screen "MTA-TiemposCmpAlta" 1280x800, template "Plantilla"
   TextField "Campo de texto_3" at 278,160 size 235x27; Text 'Tiempo apagado Sopladora'
   IOField "Campo ES_5" at 889,160 size 90x23; FormatPattern 99; Unit  min
      ProcessValue <- "TiempoSop"
   TextField "Campo de texto_1" at 278,288 size 268x27; Text 'Tiempo de compresor en vacío'
   IOField "Campo ES_1" at 889,288 size 90x23; FormatPattern 99; Unit  min
      ProcessValue <- "TiempoenVacío"
   TextField "Campo de texto_2" at 278,432 size 339x27; Text 'Tiempo sin requerimiento de compresor'
   IOField "Campo ES_2" at 889,432 size 90x23; FormatPattern 99; Unit  min
      ProcessValue <- "TiemposinReq"
   TextField "Campo de texto_4" at 286,192 size 586x36; Text 'Una vez deshabilitada una sopladora, los requisitos de marcha de compresores se mantienen durante éste tiempo.'
   TextField "Campo de texto_5" at 286,320 size 616x52; Text 'Es el tiempo máximo durante el cual el compresor quedará funcionando en vacío. Una vez cumplido éste tiempo, el compresor será pasará al estado de "sin requerimiento". Si el compresor vuelve a ser requerido en carga, se pondrá en marcha sin requerir intervención del usuario'
   TextField "Campo de texto_6" at 286,464 size 578x36; Text 'Transcurrido éste tiempo en el estado “Sin requerimiento”, pasará al estado “sin marcha”, donde sí requerirá que se pulse el botón de MARCHA en caso de ser necesitado.'
   Button "Botón_12" at 1105,638 size 160x49; TextOff 'Volver'
      on Click: function_efd93a16()
   TextField "Campo de texto_7" at 477,9 size 326x27; Text 'Configuración de Tiempos Alta presión'

screen "MTA-TorresCAV" 1280x800, template "Plantilla"
   GraphicView "Visor de gráficos_9" at 71,137 size 234x255; Picture "torreFINAL4_1"
   GraphicView "Visor de gráficos_11" at 71,137 size 234x255; Picture "torreFINAL4B_1"
   GraphicView "Visor de gráficos_14" at 71,137 size 234x255; Picture "torreFINAL4C_1"
      Visibility <- "BombaTorreON2"
   GraphicView "Visor de gráficos_1" at 271,121 size 282x311; Picture "torreFINAL4_1"
   GraphicView "Visor de gráficos_2" at 271,121 size 282x311; Picture "torreFINAL4B_1"
   GraphicView "Visor de gráficos_3" at 271,121 size 282x311; Picture "torreFINAL4C_1"
      Visibility <- "BombaTorreON2"
   Polygon "Polígono_2" at 106,411 size 18x54
      Appearance <- "FT1_AGUA"
   ScreenModuleView "Faceplate_9_2" at 831,282 size 221x68
      Guid_{11997190-23979} <- "HabilitaciónMV030"
      Guid_{11997190-23983} <- "ParadaMV030"
      Guid_{11997190-23981} <- "MarchaMV030"
      Guid_{11997190-23989} <- "SP-OFF-V030"
      Guid_{11997190-23976} <- "DeshabilitaciónMV030"
      Guid_{11997190-23987} <- "SP-ON-V030"
      Guid_{11997190-23985} <- "MenuV030"
   ScreenModuleView "Faceplate_9_1" at 831,173 size 221x68
      Guid_{11997190-23979} <- "HabilitaciónMV031"
      Guid_{11997190-23983} <- "ParadaMV031"
      Guid_{11997190-23981} <- "MarchaMV031"
      Guid_{11997190-23989} <- "SP-OFF-V031"
      Guid_{11997190-23976} <- "DeshabilitaciónMV031"
      Guid_{11997190-23987} <- "SP-ON-V031"
      Guid_{11997190-23985} <- "MenuV031"
   Polygon "Polígono_4" at 60,416 size 46x49
      Appearance <- "FT1_AGUA"
   GraphicView "Visor de gráficos_17" at 7,412 size 77x78; Picture "tuboXXX5_1"
   GraphicView "Visor de gráficos_16" at 340,421 size 190x41; Picture "tuboXXX4"
   TextField "Campo de texto_23" at 647,286 size 126x32; Text 'Ventilador 2'
   TextField "Campo de texto_3" at 647,178 size 126x32; Text 'Ventilador 1'
   GraphicIOField "Campo ES gráfico_4" at 638,358 size 511x6; PictureList "Indicador"
      ProcessValue <- "AnimaMV030"
   GraphicIOField "Campo ES gráfico_5" at 638,250 size 511x6; PictureList "Indicador"
      ProcessValue <- "AnimaMV031"
   SymbolicIOField "Campo ES simbólico_6" at 649,322 size 170x21; TextOff '0'; TextOn '1'; TextList "EstadoMotor"
      ProcessValue <- "AnimaMV030"
   SymbolicIOField "Campo ES simbólico_2" at 649,214 size 170x21; TextOff '0'; TextOn '1'; TextList "EstadoMotor"
      ProcessValue <- "AnimaMV031"
   Switch "Interruptor_5" at 782,288 size 29x29; TextOn '1'; TextOff '0'; CaptionText 'Switch'; PictureOff "A2"; PictureOn "A"
      ProcessValue <- "AutoV030"
   Switch "Interruptor_1" at 782,180 size 29x29; TextOn '1'; TextOff '0'; CaptionText 'Switch'; PictureOff "A2"; PictureOn "A"
      ProcessValue <- "AutoV031"
   GraphicIOField "Campo ES gráfico_8" at 798,700 size 418x6; PictureList "Indicador"
      ProcessValue <- "AnimaMP014"
   GraphicIOField "Campo ES gráfico_9" at 52,700 size 418x6; PictureList "Indicador"
      ProcessValue <- "AnimaMP015"
   TextField "Campo de texto_8" at 815,623 size 155x32; Text 'Backup (ESTE)'
   TextField "Campo de texto_9" at 64,623 size 182x32; Text 'Principal (OESTE)'
   SymbolicIOField "Campo ES simbólico_5" at 817,659 size 170x21; TextOff '0'; TextOn '1'; TextList "EstadoMotor"
      ProcessValue <- "AnimaMP014"
   SymbolicIOField "Campo ES simbólico_7" at 73,659 size 170x21; TextOff '0'; TextOn '1'; TextList "EstadoMotor"
      ProcessValue <- "AnimaMP015"
   GraphicView "Visor de gráficos_22" at 1067,281 size 71x70; Picture "Vent1"
   GraphicView "Visor de gráficos_23" at 1067,281 size 71x70; Picture "Vent2"
      Visibility <- "AnimaMV030"
   GraphicView "Visor de gráficos_20" at 1067,173 size 71x70; Picture "Vent1"
   GraphicView "Visor de gráficos_21" at 1067,173 size 71x70; Picture "Vent2"
      Visibility <- "AnimaMV031"
   ScreenModuleView "ControlMotor-NoAUTO_4" at 1005,625 size 203x65
      Guid_{11997190-67152} <- "DeshabilitaciónMP014"
      Guid_{11997190-67156} <- "ParadaMP014"
      Guid_{11997190-67150} <- "HabilitaciónMP014"
      Guid_{11997190-67154} <- "MarchaMP014"
   ScreenModuleView "ControlMotor-NoAUTO_5" at 259,625 size 203x65
      Guid_{11997190-67152} <- "DeshabilitaciónMP015"
      Guid_{11997190-67156} <- "ParadaMP015"
      Guid_{11997190-67150} <- "HabilitaciónMP015"
      Guid_{11997190-67154} <- "MarchaMP015"
   GraphicView "Visor de gráficos_10" at 511,450 size 13x105; Picture "tuboXXX8_1"
   GraphicView "Visor de gráficos_12" at 625,530 size 14x25; Picture "tuboXXX8_1"
   Polygon "Polígono_5" at 60,407 size 63x15
      Appearance <- "FT1_AGUA"
   TextField "Campo de texto_2" at 124,104 size 101x20; Text 'Torre 1 (NORTE)'
   TextField "Campo de texto_1" at 357,88 size 104x23; Text 'Torre 2 (SUR)'
   GraphicView "Visor de gráficos_13" at 514,528 size 125x10; Picture "Copia de tuboXXX8"
   GraphicView "Visor de gráficos_7" at 497,527 size 72x111; Picture "Bomba"
   GraphicView "Visor de gráficos_8" at 612,527 size 72x111; Picture "Bomba"
   TextField "Campo de texto_7" at 697,691 size 48x22; Text 'MP014'
   TextField "Campo de texto_6" at 582,691 size 48x22; Text 'MP015'
   TextField "Campo de texto_4" at 113,471 size 84x27; Text 'Flujostato'
   GraphicIOField "Plantilla_Campo ES gráfico_2" at 663,615 size 81x68; PictureList "Motor2"
      ProcessValue <- "AnimaMP014"
   GraphicIOField "Plantilla_Campo ES gráfico_1" at 546,615 size 81x68; PictureList "Motor2"
      ProcessValue <- "AnimaMP015"
   TextField "Campo de texto_22" at 661,479 size 90x22; Text 'Temperatura'
   IOField "Campo ES_7" at 657,499 size 98x23; FormatPattern s999999999.999; Unit  ºC
      ProcessValue <- "TempCAV"
   GraphicView "Visor de gráficos_33" at 201,338 size 118x71; Picture "tuboXXX5"
   GraphicView "Visor de gráficos_4" at 188,396 size 185x41; Picture "tuboXXX4"
   GraphicView "Visor de gráficos_5" at 108,374 size 169x37; Picture "tuboXXX4"
   GraphicView "Visor de gráficos_6" at 174,385 size 169x37; Picture "tuboXXX4"
   GraphicView "Visor de gráficos_15" at 62,386 size 130x79; Picture "tuboXXX5"
   Button "Botón_3" at 1184,68 size 48x46; TextOff '?'
      on Click: ActivateScreen("MTA-AyudaVentiladores", 0)
   TextField "Campo de texto_10" at 505,10 size 271x27; Text 'Torres de enfriamiento Cavaleto'
   GraphicIOField "Campo ES gráfico_2" at 149,135 size 76x32; PictureList "MotorTorre"
      ProcessValue <- "AnimaMV031"
   GraphicIOField "Campo ES gráfico_1" at 366,121 size 87x34; PictureList "MotorTorre"
      ProcessValue <- "AnimaMV030"

screen "MTA-TorresCH" 1280x800, template "Plantilla"
   TextField "Campo de texto_13" at 60,454 size 73x22; Text 'Presostato'
   TextField "Campo de texto_7" at 697,691 size 48x22; Text 'MP019'
   TextField "Campo de texto_6" at 582,691 size 48x22; Text 'MP018'
   GraphicView "Visor de gráficos_7" at 497,527 size 72x111; Picture "Bomba"
   GraphicView "Plantilla_Visor de gráficos_2" at 1232,6 size 35x35; Picture "ParlantesGris_1"
   GraphicView "Plantilla_Visor de gráficos_1" at 1232,6 size 35x35; Picture "ParlantesRojo"
      Visibility <- "SirenaChillers"
   GraphicView "Visor de gráficos_8" at 612,527 size 72x111; Picture "Bomba"
   Button "Botón_1" at 1220,1 size 57x44; TextOff 'Text'
      on Click: ActivateScreen("MTA-ChillersCFGSirena", 0)
   GraphicIOField "Plantilla_Campo ES gráfico_2" at 663,615 size 81x68; PictureList "Motor2"
      ProcessValue <- "AnimaciónMP019"
   GraphicIOField "Plantilla_Campo ES gráfico_1" at 546,615 size 81x68; PictureList "Motor2"
      ProcessValue <- "AnimaciónMP018"
   TextField "Campo de texto_22" at 661,479 size 90x22; Text 'Temperatura'
   Button "Botón_3" at 1184,68 size 48x46; TextOff '?'
      on Click: ActivateScreen("MTA-AyudaVentiladores", 0)
   GraphicView "Visor de gráficos_9" at 96,443 size 233x53; Picture "tuboXXX4"
   GraphicView "Visor de gráficos_11" at 62,461 size 154x79; Picture "tuboXXX5"
   GraphicView "Visor de gráficos_25" at 305,367 size 233x53; Picture "tuboXXX4"
   GraphicView "Visor de gráficos_26" at 313,379 size 233x53; Picture "tuboXXX4"
   GraphicView "Visor de gráficos_28" at 413,396 size 233x53; Picture "tuboXXX4"
   TextField "Campo de texto_10" at 511,10 size 260x27; Text 'Torres de enfriamiento Chillers'
   IOField "Campo ES_1" at 668,499 size 80x23; FormatPattern 999.99; Unit  ºC
      ProcessValue <- "TemperaturatorresCH"
   GraphicView "Visor de gráficos_1" at 271,137 size 234x255; Picture "torreFINAL4_1"
   GraphicView "Visor de gráficos_17" at 34,97 size 370x377; Picture "torreFINAL4_1"
   GraphicView "Visor de gráficos_2" at 271,137 size 234x255; Picture "torreFINAL4B_1"
   GraphicView "Visor de gráficos_5" at 34,97 size 370x377; Picture "torreFINAL4B_1"
   GraphicView "Visor de gráficos_6" at 271,137 size 234x255; Picture "torreFINAL4C_1"
      Visibility <- "BombaTorreON"
   GraphicView "Visor de gráficos_16" at 34,97 size 370x377; Picture "torreFINAL4C_1"
      Visibility <- "BombaTorreON"
   TextField "Campo de texto_2" at 364,104 size 47x20; Text 'Torre 3'
   TextField "Campo de texto_12" at 188,63 size 57x23; Text 'Torre 1'
   GraphicView "Visor de gráficos_10" at 511,530 size 13x27; Picture "tuboXXX8_1"
   Polygon "Polígono_2" at 105,487 size 18x54
      Appearance <- "Presosato"
   Polygon "Polígono_3" at 60,483 size 63x15
      Appearance <- "Presosato"
   Polygon "Polígono_4" at 59,492 size 46x49
      Appearance <- "Presosato"
   GraphicView "Visor de gráficos_12" at 625,437 size 14x117; Picture "tuboXXX8_1"
   GraphicView "Visor de gráficos_13" at 511,523 size 118x10; Picture "Copia de tuboXXX8"
   TextField "Campo de texto_1" at 589,92 size 57x23; Text 'Torre 2'
   GraphicView "Visor de gráficos_4" at 476,127 size 290x297; Picture "torreFINAL4_1"
   GraphicView "Visor de gráficos_3" at 476,127 size 290x297; Picture "torreFINAL4B_1"
   GraphicView "Visor de gráficos_15" at 476,127 size 290x297; Picture "torreFINAL4C_1"
      Visibility <- "BombaTorreON"
   ScreenModuleView "ControlMotor-NoAUTO_4" at 1021,625 size 203x65
      Guid_{11997190-67152} <- "DesMP019"
      Guid_{11997190-67156} <- "ParadaMP019"
      Guid_{11997190-67150} <- "HabMP019"
      Guid_{11997190-67154} <- "MarchaMP019"
   ScreenModuleView "ControlMotor-NoAUTO_5" at 243,625 size 203x65
      Guid_{11997190-67152} <- "DesMP018"
      Guid_{11997190-67156} <- "ParadaMP018"
      Guid_{11997190-67150} <- "HabMP018"
      Guid_{11997190-67154} <- "MarchaMP018"
   GraphicIOField "Campo ES gráfico_1" at 157,95 size 116x44; PictureList "MotorTorre"
      ProcessValue <- "AnimaciónV001"
   GraphicIOField "Campo ES gráfico_2" at 349,135 size 76x32; PictureList "MotorTorre"
      ProcessValue <- "AnimaciónV003"
   GraphicIOField "Campo ES gráfico_3" at 573,122 size 91x39; PictureList "MotorTorre"
      ProcessValue <- "AnimaciónV002"
   GraphicIOField "Campo ES gráfico_4" at 758,214 size 511x6; PictureList "Indicador"
      ProcessValue <- "AnimaciónV001"
   TextField "Campo de texto_23" at 767,142 size 126x32; Text 'Ventilador 1'
   SymbolicIOField "Campo ES simbólico_6" at 769,178 size 170x21; TextOff '0'; TextOn '1'; TextList "EstadoMotor"
      ProcessValue <- "AnimaciónV001"
   Switch "Interruptor_5" at 902,144 size 29x29; TextOn '1'; TextOff '0'; CaptionText 'Switch'; PictureOff "A2"; PictureOn "A"
      ProcessValue <- "AutoV001"
   GraphicIOField "Campo ES gráfico_5" at 758,326 size 511x6; PictureList "Indicador"
      ProcessValue <- "AnimaciónV002"
   TextField "Campo de texto_3" at 767,254 size 126x32; Text 'Ventilador 2'
   SymbolicIOField "Campo ES simbólico_2" at 769,290 size 170x21; TextOff '0'; TextOn '1'; TextList "EstadoMotor"
      ProcessValue <- "AnimaciónV002"
   Switch "Interruptor_1" at 902,256 size 29x29; TextOn '1'; TextOff '0'; CaptionText 'Switch'; PictureOff "A2"; PictureOn "A"
      ProcessValue <- "AutoV002"
   GraphicIOField "Campo ES gráfico_6" at 758,438 size 511x6; PictureList "Indicador"
      ProcessValue <- "AnimaciónV003"
   TextField "Campo de texto_4" at 767,366 size 126x32; Text 'Ventilador 3'
   SymbolicIOField "Campo ES simbólico_3" at 769,402 size 170x21; TextOff '0'; TextOn '1'; TextList "EstadoMotor"
      ProcessValue <- "AnimaciónV003"
   Switch "Interruptor_2" at 902,368 size 29x29; TextOn '1'; TextOff '0'; CaptionText 'Switch'; PictureOff "A2"; PictureOn "A"
      ProcessValue <- "AutoV003"
   TextField "Campo de texto_8" at 831,623 size 155x32; Text 'Backup (ESTE)'
   SymbolicIOField "Campo ES simbólico_5" at 833,659 size 170x21; TextOff '0'; TextOn '1'; TextList "EstadoMotor"
      ProcessValue <- "AnimaciónMP019"
   TextField "Campo de texto_9" at 47,623 size 182x32; Text 'Principal (OESTE)'
   SymbolicIOField "Campo ES simbólico_7" at 57,659 size 170x21; TextOff '0'; TextOn '1'; TextList "EstadoMotor"
      ProcessValue <- "AnimaciónMP018"
   GraphicIOField "Campo ES gráfico_8" at 814,700 size 418x6; PictureList "Indicador"
      ProcessValue <- "AnimaciónMP019"
   GraphicIOField "Campo ES gráfico_9" at 36,700 size 418x6; PictureList "Indicador"
      ProcessValue <- "AnimaciónMP018"
   ScreenModuleView "Faceplate_9_1" at 950,138 size 221x68
      Guid_{11997190-23979} <- "HabV001(1)"
      Guid_{11997190-23983} <- "ParadaV001(1)"
      Guid_{11997190-23981} <- "MarchaV001(1)"
      Guid_{11997190-23989} <- "SP-OFF-V001"
      Guid_{11997190-23976} <- "DeshV001"
      Guid_{11997190-23987} <- "SP-ON-V001"
      Guid_{11997190-23985} <- "AnimaMenuV001"
   ScreenModuleView "Faceplate_9_2" at 950,250 size 221x68
      Guid_{11997190-23979} <- "HabV002(1)"
      Guid_{11997190-23983} <- "ParadaV002(1)"
      Guid_{11997190-23981} <- "MarchaV002(1)"
      Guid_{11997190-23989} <- "SP-OFF-V002"
      Guid_{11997190-23976} <- "DeshV002"
      Guid_{11997190-23987} <- "SP-ON-V002"
      Guid_{11997190-23985} <- "AnimaMenuV002"
   ScreenModuleView "Faceplate_9_3" at 950,362 size 221x68
      Guid_{11997190-23979} <- "HabV003(1)"
      Guid_{11997190-23983} <- "ParadaV003(1)"
      Guid_{11997190-23981} <- "MarchaV003(1)"
      Guid_{11997190-23989} <- "SP-OFF-V003"
      Guid_{11997190-23976} <- "DeshV003"
      Guid_{11997190-23987} <- "SP-ON-V003"
      Guid_{11997190-23985} <- "AnimaMenuV003"
   GraphicView "Visor de gráficos_22" at 1187,137 size 71x70; Picture "Vent1"
   GraphicView "Visor de gráficos_23" at 1187,137 size 71x70; Picture "Vent2"
      Visibility <- "AnimaciónV001"
   GraphicView "Visor de gráficos_18" at 1187,360 size 71x70; Picture "Vent1"
   GraphicView "Visor de gráficos_19" at 1187,360 size 71x70; Picture "Vent2"
      Visibility <- "AnimaciónV003"
   GraphicView "Visor de gráficos_20" at 1187,249 size 71x70; Picture "Vent1"
   GraphicView "Visor de gráficos_21" at 1187,249 size 71x70; Picture "Vent2"
      Visibility <- "AnimaciónV002"
   GraphicView "Visor de gráficos_14" at 1,492 size 85x70; Picture "tuboXXX5_1"
   GraphicView "Visor de gráficos_24" at 309,399 size 237x95; Picture "tuboXXX5"

screen "SentronPAC-MTA" 1280x800, template "Plantilla"
   TextField "Campo de texto_5" at 551,10 size 179x27; Text 'Datos SENTRON PAC'
   TextField "Campo de texto_4" at 105,133 size 55x27; Text 'Actual'
   TextField "Campo de texto_6" at 337,133 size 54x27; Text 'Media'
   TextField "Campo de texto_7" at 209,133 size 68x27; Text 'Máxima'
   TextField "Campo de texto_14" at 41,165 size 16x27; Text 'R'
   IOField "Campo ES_1" at 74,165 size 110x27; FormatPattern 9999; Unit    V
      ProcessValue <- "Tension Fase R"
   IOField "Campo ES_2" at 74,197 size 110x27; FormatPattern 9999; Unit    V
      ProcessValue <- "Tension fase S"
   IOField "Campo ES_3" at 74,229 size 110x27; FormatPattern 9999; Unit    V
      ProcessValue <- "Tension Fase T"
   IOField "Campo ES_4" at 314,165 size 110x27; FormatPattern 9999; Unit    V
      ProcessValue <- "Tension Media Fase"
   IOField "Campo ES_5" at 194,165 size 110x27; FormatPattern 9999; Unit    V
      ProcessValue <- "Tension Maxima R"
   IOField "Campo ES_6" at 194,197 size 110x27; FormatPattern 9999; Unit    V
      ProcessValue <- "Tension Maxima S"
   IOField "Campo ES_7" at 194,229 size 110x27; FormatPattern 9999; Unit    V
      ProcessValue <- "Tension Maxima T"
   IOField "Campo ES_8" at 74,286 size 110x27; FormatPattern 9999; Unit    V
      ProcessValue <- "Tension Linea RS"
   IOField "Campo ES_9" at 74,318 size 110x27; FormatPattern 9999; Unit    V
      ProcessValue <- "Tension Linea ST"
   IOField "Campo ES_10" at 74,350 size 110x27; FormatPattern 9999; Unit    V
      ProcessValue <- "Tension Linea TR"
   IOField "Campo ES_11" at 314,286 size 110x27; FormatPattern 9999; Unit    V
      ProcessValue <- "Tension Media de Linea"
   IOField "Campo ES_12" at 194,286 size 110x27; FormatPattern 9999; Unit    V
      ProcessValue <- "Tension Maxima RS"
   IOField "Campo ES_13" at 194,318 size 110x27; FormatPattern 9999; Unit    V
      ProcessValue <- "Tension Maxima ST"
   IOField "Campo ES_14" at 194,350 size 110x27; FormatPattern 9999; Unit    V
      ProcessValue <- "Tension Maxima TR"
   TextField "Campo de texto_15" at 41,197 size 15x27; Text 'S'
   TextField "Campo de texto_16" at 41,229 size 15x27; Text 'T'
   TextField "Campo de texto_17" at 41,286 size 27x27; Text 'RS'
   TextField "Campo de texto_18" at 41,318 size 26x27; Text 'ST'
   TextField "Campo de texto_19" at 41,350 size 27x27; Text 'TR'
   TextField "Campo de texto_8" at 105,453 size 55x27; Text 'Actual'
   TextField "Campo de texto_9" at 337,453 size 54x27; Text 'Media'
   TextField "Campo de texto_10" at 209,453 size 68x27; Text 'Máxima'
   TextField "Campo de texto_11" at 41,485 size 16x27; Text 'R'
   TextField "Campo de texto_12" at 41,517 size 15x27; Text 'S'
   TextField "Campo de texto_13" at 41,549 size 15x27; Text 'T'
   IOField "Campo ES_15" at 74,485 size 110x27; FormatPattern 9999; Unit    A
      ProcessValue <- "Corriente fase R"
   IOField "Campo ES_16" at 74,517 size 110x27; FormatPattern 9999; Unit    A
      ProcessValue <- "Corriente Fase S"
   IOField "Campo ES_17" at 74,549 size 110x27; FormatPattern 9999; Unit    A
      ProcessValue <- "Corriente Fase T"
   IOField "Campo ES_18" at 314,485 size 110x27; FormatPattern 9999; Unit    A
      ProcessValue <- "Corriente Media"
   IOField "Campo ES_19" at 194,485 size 110x27; FormatPattern 9999; Unit    A
      ProcessValue <- "Corriente Maxima R"
   IOField "Campo ES_20" at 194,517 size 110x27; FormatPattern 9999; Unit    A
      ProcessValue <- "Corriente Maxima S"
   IOField "Campo ES_23" at 194,549 size 110x27; FormatPattern 9999; Unit    A
      ProcessValue <- "Corriente Maxima T"
   TextField "Campo de texto_20" at 719,133 size 64x27; Text 'Coseno'
   TextField "Campo de texto_21" at 703,165 size 16x27; Text 'R'
   IOField "Campo ES_24" at 725,165 size 62x27; FormatPattern 9.99; Unit    
      ProcessValue <- "Coseno R"
   TextField "Campo de texto_22" at 703,197 size 15x27; Text 'S'
   IOField "Campo ES_25" at 725,197 size 62x27; FormatPattern 9.99; Unit    
      ProcessValue <- "Coseno S"
   TextField "Campo de texto_23" at 703,229 size 15x27; Text 'T'
   IOField "Campo ES_26" at 725,229 size 62x27; FormatPattern 9.99; Unit    
      ProcessValue <- "Coseno T"
   TextField "Campo de texto_24" at 671,293 size 45x27; Text 'Total'
   IOField "Campo ES_27" at 725,293 size 62x27; FormatPattern 9.99; Unit    
      ProcessValue <- "coseno Total"
   TextField "Campo de texto_25" at 823,133 size 53x27; Text 'Activa'
   TextField "Campo de texto_26" at 942,133 size 74x27; Text 'Reactiva'
   IOField "Campo ES_28" at 797,165 size 126x27; FormatPattern 9999999; Unit  W
      ProcessValue <- "Pot.Act R"
   IOField "Campo ES_29" at 797,197 size 126x27; FormatPattern 9999999; Unit  W
      ProcessValue <- "Pot.Act S"
   IOField "Campo ES_30" at 797,229 size 126x27; FormatPattern 9999999; Unit  W
      ProcessValue <- "Pot.Act T"
   IOField "Campo ES_31" at 931,165 size 126x27; FormatPattern 9999999; Unit  var
      ProcessValue <- "Pot.ReAct R"
   IOField "Campo ES_32" at 931,197 size 126x27; FormatPattern 9999999; Unit  var
      ProcessValue <- "Pot.ReAct S"
   IOField "Campo ES_33" at 931,229 size 126x27; FormatPattern 9999999; Unit  var
      ProcessValue <- "Pot.ReAct T"
   TextField "Campo de texto_27" at 1077,133 size 80x27; Text 'Aparente'
   IOField "Campo ES_34" at 1067,165 size 121x27; FormatPattern 9999999; Unit  VA
      ProcessValue <- "Pot.ReAct R"
   IOField "Campo ES_35" at 1067,197 size 121x27; FormatPattern 9999999; Unit  VA
      ProcessValue <- "Pot.ReAct S"
   IOField "Campo ES_36" at 1067,229 size 121x27; FormatPattern 9999999; Unit  VA
      ProcessValue <- "Pot.ReAct T"
   IOField "Campo ES_21" at 797,293 size 126x27; FormatPattern 9999999; Unit  W
      ProcessValue <- "Pot Act Total"
   IOField "Campo ES_22" at 931,293 size 126x27; FormatPattern 9999999; Unit  var
      ProcessValue <- "Pot ReAct Total"
   IOField "Campo ES_37" at 1067,293 size 121x27; FormatPattern 9999999; Unit  VA
      ProcessValue <- "Pot Apa Total"
   TextField "Campo de texto_30" at 695,461 size 95x27; Text 'Frecuencia'
   TextField "Campo de texto_31" at 695,493 size 171x27; Text 'Desbalance Tensión'
   TextField "Campo de texto_32" at 695,525 size 182x27; Text 'Desbalance Corriente'
   IOField "Campo ES_38" at 893,461 size 110x27; FormatPattern 99.99; Unit    Hz
      ProcessValue <- "Frecuencia"
   IOField "Campo ES_39" at 893,493 size 110x27; FormatPattern 99.99; Unit    %
      ProcessValue <- "desbalance de tension"
   IOField "Campo ES_40" at 893,525 size 110x27; FormatPattern 99.99; Unit    %
      ProcessValue <- "desbalance de corriente"
   TextField "Campo de texto_29" at 465,133 size 41x27; Text 'THD'
   TextField "Campo de texto_33" at 465,453 size 41x27; Text 'THD'
   IOField "Campo ES_41" at 434,165 size 110x27; FormatPattern 99.999; Unit    %
      ProcessValue <- "THD-R TensionFase R"
   IOField "Campo ES_42" at 434,197 size 110x27; FormatPattern 99.999; Unit    %
      ProcessValue <- "THD-R Tension Fase S"
   IOField "Campo ES_43" at 434,229 size 110x27; FormatPattern 99.999; Unit    %
      ProcessValue <- "THD-R Tension Fase T"
   IOField "Campo ES_47" at 434,485 size 110x27; FormatPattern 99.999; Unit    %
      ProcessValue <- "THD-R Corriente Fase R"
   IOField "Campo ES_48" at 434,517 size 110x27; FormatPattern 99.999; Unit    %
      ProcessValue <- "THD-R Corriente Fase S"
   IOField "Campo ES_49" at 434,549 size 110x27; FormatPattern 99.999; Unit    %
      ProcessValue <- "THD-R Corriente Fase T"
   TextField "Campo de texto_34" at 31,100 size 603x27; Text 'Tensión'
   TextField "Campo de texto_35" at 31,420 size 603x27; Text 'Corriente'
   TextField "Campo de texto_1" at 650,100 size 609x27; Text 'Potencia'
   TextField "Campo de texto_2" at 655,420 size 601x27; Text 'General'
   Button "Botón_1" at 565,186 size 50x49; TextOff 'Text'; PictureOff "Gráfico_8"
      on Press: ActivateScreen("Graf-Fase", 0)
   Button "Botón_2" at 565,315 size 50x49; TextOff 'Text'; PictureOff "Gráfico_8"
      on Press: ActivateScreen("Graf-Linea", 0)
   Button "Botón_3" at 565,506 size 50x49; TextOff 'Text'; PictureOff "Gráfico_8"
      on Press: ActivateScreen("Graf-Corrientes", 0)
   Button "Botón_4" at 1197,186 size 50x49; TextOff 'Text'; PictureOff "Gráfico_8"
      on Press: ActivateScreen("Graf-Pot", 0)
   Button "Botón_5" at 1197,282 size 50x49; TextOff 'Text'; PictureOff "Gráfico_8"
      on Press: ActivateScreen("Graf-PotTotal", 0)

screen "MTA-AyudaCmpBaja" 1280x800, template "Plantilla"
   GraphicIOField "Campo ES gráfico_7" at 279,380 size 178x52; PictureList "BaseSullChico"
      ProcessValue <- "UNO"
   GraphicIOField "Campo ES gráfico_1" at 351,380 size 178x52; PictureList "BaseSullChico"
      ProcessValue <- "UNO"
   GraphicView "Visor de gráficos_3" at 269,294 size 269x127; Picture "baja2X_2"
   GraphicView "Visor de gráficos_9" at 335,168 size 269x127; Picture "baja2Xd_1"
   TextField "Campo de texto_11" at 50,259 size 199x76; Text 'El modo local transfiere el control del Compresor a su panel original'
   TextField "Campo de texto_12" at 39,229 size 210x42; Text 'Activación de modo "LOCAL"'
   TextField "Campo de texto_2" at 145,116 size 210x42; Text 'Indicación de modo "LOCAL"'
   TextField "Campo de texto_8" at 762,110 size 352x94; Text 'La Deshabilitación del Compresor provoca también la detención del mismo. La Habilitación del Compresor permite su operaración desde el panel.'
   TextField "Campo de texto_9" at 946,227 size 230x76; Text 'Para poder marchar el Compresor es necesario que el mismo esté habilitado'
   TextField "Campo de texto_4" at 751,85 size 203x42; Text 'Habilitación/Deshabilitación'
   TextField "Campo de texto_13" at 991,455 size 195x42; Text 'Orden de Parar Compresor'
   GraphicView "Visor de gráficos_5" at 920,329 size 202x77; Picture "menu2"
   GraphicIOField "Campo ES gráfico_2" at 621,403 size 507x6; PictureList "Indicador"
      ProcessValue <- "UNO"
   TextField "Campo de texto_14" at 589,454 size 160x42; Text 'Estado del Compresor'
   TextField "Campo de texto_15" at 615,261 size 108x61; Text 'Nombre del Compresor'
   GraphicView "Visor de gráficos_1" at 804,336 size 31x31; Picture "A2"
   TextField "Campo de texto_1" at 789,269 size 54x42; Text 'Manual'
   TextField "Campo de texto_16" at 335,457 size 134x42; Text 'Código de Colores'
   GraphicView "Visor de gráficos_4" at 920,497 size 202x77; Picture "menu5"
   GraphicIOField "Campo ES gráfico_3" at 621,571 size 507x6; PictureList "Indicador"
      ProcessValue <- "UNO"
   GraphicView "Visor de gráficos_2" at 806,505 size 31x31; Picture "A"
   TextField "Campo de texto_17" at 798,443 size 38x42; Text 'Auto'
   TextField "Campo de texto_6" at 477,590 size 726x99; Text 'Modo Automático Cada Compresor se pondrá en Marcha si la Presión de línea sensada se encuentra por debajo del valor de "On" y se apagará una vez superado el valor de "Off" El Compresor mantiene su marcha 5 minutos después de haber superado el valor de "Off" para evitar arranques consecutivos del mismo.'
   TextField "Campo de texto_5" at 29,520 size 471x213; Text 'El funcionamiento descripto solo se aplica a los compresores: ATLAS 2 ATLAS 3 SULLAIR 0 SULLAIR 1 El Compresor SULLAIR2 NO PUEDE SER CONTROLADO DESDE EL PANEL'
   TextField "Campo de texto_10" at 529,9 size 246x27; Text 'Ayuda: Compresores de Baja'
   TextField "Campo de texto_7" at 645,334 size 116x39; Text 'Sullair 0'
   SymbolicIOField "Campo ES simbólico_7" at 647,370 size 242x21; TextOff '0'; TextOn '1'; TextList "EstadoMotor"
      ProcessValue <- "UNO"
   TextField "Campo de texto_3" at 645,502 size 116x39; Text 'Sullair 0'
   SymbolicIOField "Campo ES simbólico_1" at 647,538 size 242x21; TextOff '0'; TextOn '1'; TextList "EstadoMotor"
      ProcessValue <- "UNO"
   Switch "Interruptor_6" at 267,305 size 40x40; TextOn '1'; TextOff '0'; CaptionText 'Switch'; PictureOff "MECH2"; PictureOn "MECH1"
      ProcessValue <- "MantM062"

screen "MTA-CompALTA" 1280x800, template "Plantilla"
   GraphicIOField "Plantilla_Campo ES gráfico_3" at 758,425 size 65x60; PictureList "Motor2"
      ProcessValue <- "AnimMotorMC001"
   GraphicIOField "Plantilla_Campo ES gráfico_4" at 685,353 size 65x60; PictureList "Motor2"
      ProcessValue <- "AnimMotorMC002"
   GraphicIOField "Plantilla_Campo ES gráfico_5" at 612,281 size 65x60; PictureList "Motor2"
      ProcessValue <- "AnimMotorMC004"
   GraphicIOField "Plantilla_Campo ES gráfico_2" at 539,209 size 65x60; PictureList "Motor2"
      ProcessValue <- "AnimMotorMC005"
   GraphicView "Visor de gráficos_2" at 492,46 size 254x172; Picture "bell1"
   GraphicView "Visor de gráficos_18" at 492,46 size 254x172; Picture "Beliss2_1"
      Visibility <- "MantMC003"
   GraphicIOField "Plantilla_Campo ES gráfico_1" at 490,113 size 100x102; PictureList "MotorBelliss"
      ProcessValue <- "AnimMotorMC003"
   GraphicView "Visor de gráficos_3" at 569,134 size 246x148; Picture "ALTA1_1"
   ScreenModuleView "Faceplate_8_1" at 781,145 size 47x30
      Guid_{11997190-23981} <- "EV3"
   GraphicView "Visor de gráficos_8" at 1175,577 size 29x50; Picture "Gráfico_2"
   GraphicView "Visor de gráficos_7" at 885,605 size 391x113; Picture "tanque1X2"
   TextField "Plantilla_Campo de texto_1" at 1141,578 size 32x23; Text 'PT2'
   IOField "Campo ES_1" at 943,632 size 108x28; FormatPattern s999.9; Unit   bar
      ProcessValue <- "PresiónALTA"
   Button "Botón_7" at 1119,186 size 128x41; TextOff 'Tiempos'
      on Click: ActivateScreen("MTA-TiemposCmpAlta", 0)
   Button "Botón_12" at 1119,234 size 128x41; TextOff 'Presiones'
      on Click: ActivateScreen("MTA-CFGALTA", 0)
   Button "Botón_13" at 1119,138 size 128x41; TextOff 'Sopladoras'
      on Click: ActivateScreen("MTA-Sopladoras", 0)
   Button "Botón_14" at 641,627 size 160x46; TextOff 'CFG Avisos'
      on Click: ActivateScreen("MTA-CFGAvisosALTA", 0)
   TextField "Campo de texto_2" at 519,9 size 242x27; Text 'Compresores de Alta Presión'
   ScreenModuleView "Faceplate_8_5" at 927,289 size 47x30
      Guid_{11997190-23981} <- "EV4"
   ScreenModuleView "Faceplate_8_4" at 1000,361 size 47x30
      Guid_{11997190-23981} <- "EV2"
   GraphicView "Visor de gráficos_19" at 569,134 size 246x148; Picture "LOCAl"
      Visibility <- "MantMC005"
   ScreenModuleView "Faceplate_8_2" at 854,217 size 47x30
      Guid_{11997190-23981} <- "EV5"
   GraphicView "Visor de gráficos_4" at 642,206 size 246x148; Picture "ALTA1_3"
   GraphicView "Visor de gráficos_22" at 642,206 size 246x148; Picture "LOCAl"
      Visibility <- "MantMC004"
   GraphicView "Visor de gráficos_5" at 715,278 size 246x148; Picture "ALTA1_3"
   GraphicView "Visor de gráficos_21" at 715,278 size 246x148; Picture "LOCAl"
      Visibility <- "MantMC002"
   GraphicView "Visor de gráficos_6" at 788,350 size 246x148; Picture "ALTA1_3"
   GraphicView "Visor de gráficos_20" at 788,350 size 246x148; Picture "LOCAl"
      Visibility <- "MantMC001"
   ScreenModuleView "Faceplate_8_3" at 1072,433 size 47x30
      Guid_{11997190-23981} <- "EV1"
   ScreenModuleView "Faceplate_8_6" at 748,113 size 47x30
      Guid_{11997190-23981} <- "EV3b"
   Button "Botón_3" at 1181,68 size 48x46; TextOff '?'
      on Click: ActivateScreen("MTA-AyudaCmpAlta", 0)
   ScreenModuleView "Faceplate_8_7" at 1144,505 size 47x30
      Guid_{11997190-23981} <- "EV6"
   GraphicIOField "Plantilla_Campo ES gráfico_6" at 831,497 size 65x60; PictureList "Motor2"
      ProcessValue <- "AnimMotorMC006"
   GraphicView "Visor de gráficos_1" at 861,422 size 246x148; Picture "ALTA1_3"
   GraphicView "Visor de gráficos_9" at 861,422 size 246x148; Picture "LOCAl"
      Visibility <- "MantMC006"
   GraphicIOField "Campo ES gráfico_4" at 6,182 size 374x6; PictureList "Indicador"
      ProcessValue <- "AnimMotorMC003"
   SymbolicIOField "Campo ES simbólico_4" at 25,154 size 178x21; TextOff '0'; TextOn '1'; TextList "EstadoMotor"
      ProcessValue <- "AnimMotorMC003"
   TextField "Campo de texto_1" at 19,121 size 55x32; Text 'Bellis'
   GraphicIOField "Campo ES gráfico_5" at 118,341 size 374x6; PictureList "Indicador"
      ProcessValue <- "AnimMotorMC004"
   TextField "Campo de texto_6" at 127,280 size 67x32; Text 'ABC-4'
   SymbolicIOField "Campo ES simbólico_5" at 137,313 size 186x21; TextOff '0'; TextOn '1'; TextList "EstadoMotor"
      ProcessValue <- "AnimMotorMC004"
   GraphicIOField "Campo ES gráfico_1" at 191,422 size 374x6; PictureList "Indicador"
      ProcessValue <- "AnimMotorMC002"
   TextField "Campo de texto_8" at 200,361 size 67x32; Text 'ABC-3'
   SymbolicIOField "Campo ES simbólico_1" at 210,394 size 186x21; TextOff '0'; TextOn '1'; TextList "EstadoMotor"
      ProcessValue <- "AnimMotorMC002"
   GraphicIOField "Campo ES gráfico_3" at 44,262 size 373x6; PictureList "Indicador"
      ProcessValue <- "AnimMotorMC005"
   TextField "Campo de texto_10" at 53,201 size 67x32; Text 'ABC-5'
   SymbolicIOField "Campo ES simbólico_3" at 63,234 size 194x21; TextOff '0'; TextOn '1'; TextList "EstadoMotor"
      ProcessValue <- "AnimMotorMC005"
   GraphicIOField "Campo ES gráfico_2" at 264,502 size 374x6; PictureList "Indicador"
      ProcessValue <- "AnimMotorMC001"
   TextField "Campo de texto_9" at 273,441 size 67x32; Text 'ABC-2'
   SymbolicIOField "Campo ES simbólico_2" at 283,474 size 186x21; TextOff '0'; TextOn '1'; TextList "EstadoMotor"
      ProcessValue <- "AnimMotorMC001"
   GraphicIOField "Campo ES gráfico_16" at 337,582 size 374x6; PictureList "Indicador"
      ProcessValue <- "AnimMotorMC006"
   TextField "Campo de texto_3" at 346,521 size 67x32; Text 'ABC-1'
   SymbolicIOField "Campo ES simbólico_11" at 356,554 size 186x21; TextOff '0'; TextOn '1'; TextList "EstadoMotor"
      ProcessValue <- "AnimMotorMC006"
   IOField "Campo ES_6" at 255,157 size 85x19; FormatPattern 999999999; Unit  hs
      ProcessValue <- "HORAS3"
      Appearance <- "EstadoMantMC003"
   IOField "Campo ES_2" at 367,316 size 85x19; FormatPattern 999999999; Unit  hs
      ProcessValue <- "HORAS4"
      Appearance <- "EstadoMantMC004"
   IOField "Campo ES_3" at 439,397 size 85x19; FormatPattern 999999999; Unit  hs
      ProcessValue <- "HORAS2"
      Appearance <- "EstadoMantMC002"
   IOField "Campo ES_5" at 292,237 size 85x19; FormatPattern 999999999; Unit  hs
      ProcessValue <- "HORAS5"
      Appearance <- "EstadoMantMC005"
   IOField "Campo ES_4" at 512,477 size 85x19; FormatPattern 999999999; Unit  hs
      ProcessValue <- "HORAS1"
      Appearance <- "EstadoMantMC001"
   IOField "Campo ES_7" at 585,557 size 85x19; FormatPattern 999999999; Unit  hs
      ProcessValue <- "HORAS6"
      Appearance <- "EstadoMantMC006"
   ScreenModuleView "Faceplate_6_1" at 283,125 size 57x28; ScreenModuleType ""
      Guid_{11997190-52606} <- "IndV3"
      Guid_{11997190-52610} <- "IndR3"
      Guid_{11997190-52608} <- "IndVparp3"
   ScreenModuleView "Faceplate_6_5" at 395,284 size 57x28; ScreenModuleType ""
      Guid_{11997190-52606} <- "IndV4"
      Guid_{11997190-52610} <- "IndR4"
      Guid_{11997190-52608} <- "IndVparp4"
   ScreenModuleView "Faceplate_6_4" at 468,365 size 57x28; ScreenModuleType ""
      Guid_{11997190-52606} <- "IndV2"
      Guid_{11997190-52610} <- "IndR2"
      Guid_{11997190-52608} <- "IndVparp2"
   ScreenModuleView "Faceplate_6_2" at 321,205 size 57x28; ScreenModuleType ""
      Guid_{11997190-52606} <- "IndV5"
      Guid_{11997190-52610} <- "IndR5"
      Guid_{11997190-52608} <- "IndVparp5"
   ScreenModuleView "Faceplate_6_3" at 541,445 size 57x28; ScreenModuleType ""
      Guid_{11997190-52606} <- "IndV1"
      Guid_{11997190-52610} <- "IndR1"
      Guid_{11997190-52608} <- "IndVparp1"
   GraphicIOField "Campo ES gráfico_6" at 348,125 size 9x45; PictureList "BarraPrioridades"
      ProcessValue <- "VCMP3"
      Visibility <- "MantMC003"
   GraphicIOField "Campo ES gráfico_9" at 357,125 size 9x45; PictureList "BarraPrioridades_1"
      ProcessValue <- "PriRealCMP3"
      Visibility <- "MantMC003"
   SymbolicIOField "Campo ES simbólico_6" at 86,124 size 160x29; TextOff '0'; TextOn '1'; TextList "EstadoCmpAlta"
      ProcessValue <- "Est3"
      Visibility <- "MantMC003"
   Button "Botón_11" at 6,116 size 374x64; TextOff 'Text'
      on Click: ActivateScreen("MTA-ALTAMC003", 0)
   Switch "Interruptor_1" at 250,125 size 29x29; TextOn '1'; TextOff '0'; CaptionText 'Switch'; PictureOff "A2"; Authorization "Operación"; PictureOn "A"
      ProcessValue <- "Auto3"
      Visibility <- "MantMC003"
   Switch "Interruptor_10" at 863,114 size 40x40; TextOn '1'; TextOff '0'; CaptionText 'Switch'; PictureOff "MECH2"; Authorization "Operación"; PictureOn "MECH1"
      ProcessValue <- "MantMC003"
   GraphicIOField "Campo ES gráfico_14" at 459,286 size 9x45; PictureList "BarraPrioridades"
      ProcessValue <- "VCMP4"
      Visibility <- "MantMC004"
   GraphicIOField "Campo ES gráfico_15" at 468,286 size 9x45; PictureList "BarraPrioridades_1"
      ProcessValue <- "PriRealCMP4"
      Visibility <- "MantMC004"
   SymbolicIOField "Campo ES simbólico_10" at 195,283 size 160x29; TextOff '0'; TextOn '1'; TextList "EstadoCmpAlta"
      ProcessValue <- "Est4"
      Visibility <- "MantMC004"
   Button "Botón_6" at 118,275 size 374x64; TextOff 'Text'
      on Click: ActivateScreen("MTA-ALTAMC004", 0)
   Switch "Interruptor_5" at 360,285 size 29x29; TextOn '1'; TextOff '0'; CaptionText 'Switch'; PictureOff "A2"; Authorization "Operación"; PictureOn "A"
      ProcessValue <- "Auto4"
      Visibility <- "MantMC004"
   Switch "Interruptor_9" at 1009,258 size 40x40; TextOn '1'; TextOff '0'; CaptionText 'Switch'; PictureOff "MECH2"; Authorization "Operación"; PictureOn "MECH1"
      ProcessValue <- "MantMC004"
   GraphicIOField "Campo ES gráfico_12" at 532,367 size 9x45; PictureList "BarraPrioridades"
      ProcessValue <- "VCMP2"
      Visibility <- "MantMC002"
   GraphicIOField "Campo ES gráfico_13" at 541,367 size 9x45; PictureList "BarraPrioridades_1"
      ProcessValue <- "PriRealCMP2"
      Visibility <- "MantMC002"
   SymbolicIOField "Campo ES simbólico_9" at 269,364 size 160x29; TextOff '0'; TextOn '1'; TextList "EstadoCmpAlta"
      ProcessValue <- "Est2"
      Visibility <- "MantMC002"
   Button "Botón_8" at 191,356 size 374x64; TextOff 'Text'
      on Click: ActivateScreen("MTA-ALTAMC002", 0)
   Switch "Interruptor_4" at 433,366 size 29x29; TextOn '1'; TextOff '0'; CaptionText 'Switch'; PictureOff "A2"; Authorization "Operación"; PictureOn "A"
      ProcessValue <- "Auto2"
      Visibility <- "MantMC002"
   Switch "Interruptor_8" at 1082,330 size 40x40; TextOn '1'; TextOff '0'; CaptionText 'Switch'; PictureOff "MECH2"; Authorization "Operación"; PictureOn "MECH1"
      ProcessValue <- "MantMC002"
   GraphicIOField "Campo ES gráfico_7" at 385,207 size 9x45; PictureList "BarraPrioridades"
      ProcessValue <- "VCMP5"
      Visibility <- "MantMC005"
   GraphicIOField "Campo ES gráfico_10" at 394,207 size 9x45; PictureList "BarraPrioridades_1"
      ProcessValue <- "PriRealCMP5"
      Visibility <- "MantMC005"
   SymbolicIOField "Campo ES simbólico_7" at 120,204 size 160x29; TextOff '0'; TextOn '1'; TextList "EstadoCmpAlta"
      ProcessValue <- "Est5"
      Visibility <- "MantMC005"
   Switch "Interruptor_6" at 936,186 size 40x40; TextOn '1'; TextOff '0'; CaptionText 'Switch'; PictureOff "MECH2"; Authorization "Operación"; PictureOn "MECH1"
      ProcessValue <- "MantMC005"
   GraphicIOField "Campo ES gráfico_8" at 605,447 size 9x45; PictureList "BarraPrioridades"
      ProcessValue <- "VCMP1"
      Visibility <- "MantMC001"
   GraphicIOField "Campo ES gráfico_11" at 614,447 size 9x45; PictureList "BarraPrioridades_1"
      ProcessValue <- "PriRealCMP1"
      Visibility <- "MantMC001"
   SymbolicIOField "Campo ES simbólico_8" at 341,444 size 160x29; TextOff '0'; TextOn '1'; TextList "EstadoCmpAlta"
      ProcessValue <- "Est1"
      Visibility <- "MantMC001"
   Button "Botón_9" at 264,436 size 374x64; TextOff 'Text'
      on Click: ActivateScreen("MTA-ALTAMC001", 0)
   Switch "Interruptor_3" at 504,445 size 29x29; TextOn '1'; TextOff '0'; CaptionText 'Switch'; PictureOff "A2"; Authorization "Operación"; PictureOn "A"
      ProcessValue <- "Auto1"
      Visibility <- "MantMC001"
   Switch "Interruptor_7" at 1155,402 size 40x40; TextOn '1'; TextOff '0'; CaptionText 'Switch'; PictureOff "MECH2"; Authorization "Operación"; PictureOn "MECH1"
      ProcessValue <- "MantMC001"
   Switch "Interruptor_11" at 1228,474 size 40x40; TextOn '1'; TextOff '0'; CaptionText 'Switch'; PictureOff "MECH2"; Authorization "Operación"; PictureOn "MECH1"
      ProcessValue <- "MantMC006"
   ScreenModuleView "Faceplate_6_6" at 614,525 size 57x28; ScreenModuleType ""
      Guid_{11997190-52606} <- "IndV6"
      Guid_{11997190-52610} <- "IndR6"
      Guid_{11997190-52608} <- "IndVparp6"
   GraphicIOField "Campo ES gráfico_17" at 678,527 size 9x45; PictureList "BarraPrioridades"
      ProcessValue <- "VCMP6"
      Visibility <- "MantMC001"
   GraphicIOField "Campo ES gráfico_18" at 687,527 size 9x45; PictureList "BarraPrioridades_1"
      ProcessValue <- "PriRealCMP6"
      Visibility <- "MantMC001"
   SymbolicIOField "Campo ES simbólico_12" at 414,524 size 160x29; TextOff '0'; TextOn '1'; TextList "EstadoCmpAlta"
      ProcessValue <- "Est6"
      Visibility <- "MantMC001"
   Button "Botón_1" at 337,516 size 374x64; TextOff 'Text'
      on Click: ActivateScreen("MTA-ALTAMC006", 0)
   Switch "Interruptor_12" at 577,525 size 29x29; TextOn '1'; TextOff '0'; CaptionText 'Switch'; PictureOff "A2"; Authorization "Operación"; PictureOn "A"
      ProcessValue <- "Auto6"
      Visibility <- "MantMC001"
   Button "Botón_10" at 45,196 size 374x64; TextOff 'Text'
      on Click: ActivateScreen("MTA-ALTAMC005", 0)
   Switch "Interruptor_2" at 284,206 size 29x29; TextOn '1'; TextOff '0'; CaptionText 'Switch'; PictureOff "A2"; Authorization "Operación"; PictureOn "A"
      ProcessValue <- "Auto5"
      Visibility <- "MantMC005"
   Rectangle "Rectángulo_22" at 20,556 size 225x82
      Visibility <- "DB_ALA_MEM_x199"
      Appearance <- "DB_ALA_MEM_x199"
   TextField "Campo de texto_4" at 27,564 size 212x67; Text 'Falla por relé de frecuencia Reconocer alarma'
      Visibility <- "DB_ALA_MEM_x199"
   IOField "Campo ES_8" at 83,495 size 96x32; FormatPattern 1
      ProcessValue <- "DB_ALA_MEM_x199"

screen "MTA-ALTAMC006" 1280x800, template "Plantilla-Alta-Cmp"
   Button "Botón_1" at 186,441 size 48x38; TextOff 'Incrementar'; Authorization "Operación"; PictureOff "Gráfico_3"
      on Press: SetBit("IncP6")
      on Release: ResetBit("IncP6")
   Button "Botón_2" at 186,401 size 48x38; TextOff 'Decrementar'; Authorization "Operación"; PictureOff "Gráfico_1"
      on Press: SetBit("DecP6")
      on Release: ResetBit("DecP6")
   Button "Botón_7" at 390,106 size 40x38; TextOff 'Text'; PictureOff "x"
      on Click: function_efd93a16()
   Button "Botón_8" at 306,600 size 96x35; TextOff 'Hecho'; Authorization "Administración de usuarios"
      on Press: SetTag("Varios_UltimoMantMC006_1", "HORAS6")
   TextField "Campo de texto_6" at 266,362 size 72x27; Text 'Seteada'
   TextField "Campo de texto_7" at 82,426 size 84x27; Text 'Prioridad'
   TextField "Campo de texto_8" at 362,363 size 40x27; Text 'Real'
   TextField "Campo de texto_11" at 26,343 size 158x27; Text 'Seteo de Prioridad'
   GraphicIOField "Campo ES gráfico_3" at 294,402 size 16x78; PictureList "BarraPrioridades"
      ProcessValue <- "VCMP6"
   GraphicIOField "Campo ES gráfico_5" at 374,402 size 16x78; PictureList "BarraPrioridades_1"
      ProcessValue <- "PriRealCMP6"
   SymbolicIOField "Campo ES simbólico_2" at 9,290 size 424x37; TextOff '0'; TextOn '1'; TextList "EstadoCmpAlta"
      ProcessValue <- "Est6"
      Visibility <- "MantMC006"
   TextField "Campo de texto_16" at 521,10 size 279x27; Text 'Menú Compresor ABC-1 (MC006)'
   TextField "Campo de texto_1" at 32,510 size 326x27; Text 'Tiempo de funcionamiento acumulado'
   TextField "Campo de texto_4" at 32,570 size 231x27; Text 'Próximo mantenimiento #1'
   TextField "Campo de texto_5" at 32,635 size 231x27; Text 'Próximo mantenimiento #2'
   Button "Botón_3" at 306,665 size 96x35; TextOff 'Hecho'; Authorization "Administración de usuarios"
      on Press: SetTag("Varios_UltimoMantMC006_2", "HORAS6")
   IOField "Campo ES_4" at 574,609 size 96x32; FormatPattern 99; Unit  min
      ProcessValue <- "DB-PurgaComAlta_Toff_PurgaABC1"
   IOField "Campo ES_5" at 574,654 size 96x32; FormatPattern 99; Unit  seg
      ProcessValue <- "DB-PurgaComAlta_Ton_PurgaABC1"
   TextField "Campo de texto_2" at 459,613 size 97x27; Text 'Tiempo Off'
   TextField "Campo de texto_3" at 459,655 size 96x27; Text 'Tiempo On'
   Switch "Interruptor_2" at 459,548 size 120x40; TextOff 'OFF'; TextOn 'ON'; CaptionText 'Switch'
      ProcessValue <- "DB-PurgaComAlta_Habil_PurgaABC1"
   Button "Botón_4" at 595,548 size 80x40; TextOff 'Prueba'
      on Press: SetBit("DB-PurgaComAlta_Prueba_PurgaABC1")
      on Release: ResetBit("DB-PurgaComAlta_Prueba_PurgaABC1")
      ObjectEnable <- "MC006_EVP"
      Appearance <- "MC006_EVP"
   TextField "Campo de texto_9" at 456,510 size 131x27; Text 'Ciclo de Purga:'
   GraphicIOField "Campo ES gráfico_2" at 10,280 size 422x6; PictureList "Indicador"
      ProcessValue <- "AnimMotorMC006"
   SymbolicIOField "Campo ES simbólico_4" at 19,246 size 290x21; TextOff '0'; TextOn '1'; TextList "EstadoMotor"
      ProcessValue <- "AnimMotorMC006"
   Button "Botón_6" at 13,154 size 88x62; TextOff 'ABC 1'
   Switch "Interruptor_1" at 150,167 size 37x37; TextOn '1'; TextOff '0'; CaptionText 'Switch'; PictureOff "A2"; Authorization "Operación"; PictureOn "A"
      ProcessValue <- "Auto6"
      Visibility <- "MantMC006"
   ScreenModuleView "Faceplate_6_1" at 342,236 size 76x34; ScreenModuleType ""
      Guid_{11997190-52606} <- "IndV6"
      Guid_{11997190-52610} <- "IndR6"
      Guid_{11997190-52608} <- "IndVparp6"
   ScreenModuleView "Faceplate_7_1" at 213,158 size 207x70
      Guid_{11997190-23983} <- "ParadaMC006"
      Guid_{11997190-90325} <- "MarchaMC006"
      Guid_{11997190-23981} <- "MarchaMC006"
      Guid_{11997190-89805} <- "SPONF6"
      Guid_{11997190-180841} <- "MantMC006"
      Guid_{11997190-89807} <- "SPOFFF6"
      Guid_{11997190-89795} <- "ForzandoMarcha6"
      Guid_{11997190-90329} <- "ForzarParada6"
      Guid_{11997190-88662} <- "MarchaOK6"
      Guid_{11997190-23985} <- "AnimMenuMC006"
   IOField "Campo ES_7" at 20,535 size 173x35; Authorization "Administración de usuarios"; FormatPattern 999999999; Unit  hs
      ProcessValue <- "HORAS6"
      Appearance <- "EstadoMantMC006"
   IOField "Campo ES_1" at 200,535 size 80x35; Authorization "Administración de usuarios"; FormatPattern 99; Unit  min
      ProcessValue <- "MIN6"
   IOField "Campo ES_2" at 20,595 size 173x35; FormatPattern 999999999; Unit  hs
      ProcessValue <- "ProxMantMC006_1"
      Appearance <- "LimiteMantMC006_1"
   IOField "Campo ES_3" at 20,660 size 173x35; FormatPattern 999999999; Unit  hs
      ProcessValue <- "ProxMantMC006_2"
      Appearance <- "LimiteMantMC006_2"